// TIA Portal project "Sistema_de_silos" (V16) (continued)
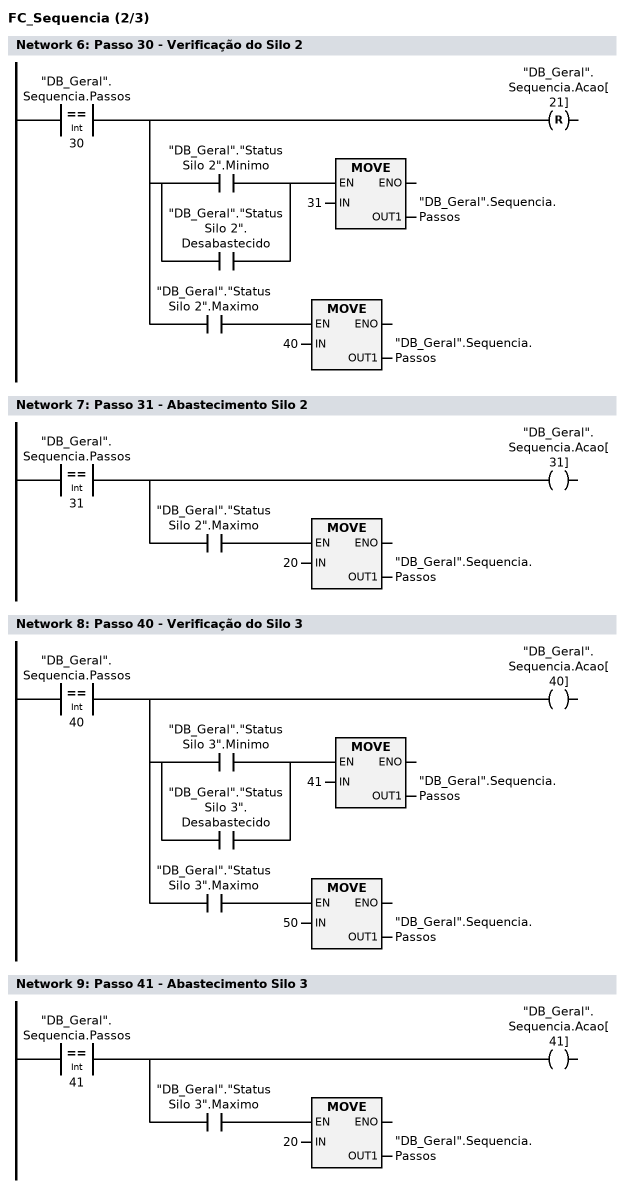
   RUNG wire#powerrail
      { S7_Templates := "SrcType := Int" } EQ_Contact(in1 := "DB_Geral".Sequencia.Passos, in2 := 30)
      wire#w1
      R_Coil( "DB_Geral".Sequencia.Acao[21] )
   END_RUNG
   RUNG wire#w1
      Contact( "DB_Geral"."Status Silo 2".Minimo )
      wire#w2
      Move(in := 31, out1 => "DB_Geral".Sequencia.Passos)
   END_RUNG
   RUNG wire#w1
      Contact( "DB_Geral"."Status Silo 2".Desabastecido )
   END_RUNG wire#w2
   RUNG wire#w1
      Contact( "DB_Geral"."Status Silo 2".Maximo )
      Move(in := 40, out1 => "DB_Geral".Sequencia.Passos)
   END_RUNG
   // the same network as SCL:
   #_w1 := "DB_Geral".Sequencia.Passos = 30;
   IF #_w1 THEN "DB_Geral".Sequencia.Acao[21] := FALSE; END_IF;
   IF #_w1 AND ("DB_Geral"."Status Silo 2".Minimo OR "DB_Geral"."Status Silo 2".Desabastecido) THEN
       "DB_Geral".Sequencia.Passos := 31;
   END_IF;
   IF #_w1 AND "DB_Geral"."Status Silo 2".Maximo THEN "DB_Geral".Sequencia.Passos := 40; END_IF;
END_REGION

REGION Network 7: Passo 31 - Abastecimento Silo 2
   RUNG wire#powerrail
      { S7_Templates := "SrcType := Int" } EQ_Contact(in1 := "DB_Geral".Sequencia.Passos, in2 := 31)
      wire#w1
      Coil( "DB_Geral".Sequencia.Acao[31] )
   END_RUNG
   RUNG wire#w1
      Contact( "DB_Geral"."Status Silo 2".Maximo )
      Move(in := 20, out1 => "DB_Geral".Sequencia.Passos)
   END_RUNG
   // the same network as SCL:
   "DB_Geral".Sequencia.Acao[31] := "DB_Geral".Sequencia.Passos = 31;
   IF ("DB_Geral".Sequencia.Passos = 31) AND "DB_Geral"."Status Silo 2".Maximo THEN
       "DB_Geral".Sequencia.Passos := 20;
   END_IF;
END_REGION

REGION Network 8: Passo 40 - Verificação do Silo 3
   RUNG wire#powerrail
      { S7_Templates := "SrcType := Int" } EQ_Contact(in1 := "DB_Geral".Sequencia.Passos, in2 := 40)
      wire#w1
      Coil( "DB_Geral".Sequencia.Acao[40] )
   END_RUNG
   RUNG wire#w1
      Contact( "DB_Geral"."Status Silo 3".Minimo )
      wire#w2
      Move(in := 41, out1 => "DB_Geral".Sequencia.Passos)
   END_RUNG
   RUNG wire#w1
      Contact( "DB_Geral"."Status Silo 3".Desabastecido )
   END_RUNG wire#w2
   RUNG wire#w1
      Contact( "DB_Geral"."Status Silo 3".Maximo )
      Move(in := 50, out1 => "DB_Geral".Sequencia.Passos)
   END_RUNG
   // the same network as SCL:
   "DB_Geral".Sequencia.Acao[40] := "DB_Geral".Sequencia.Passos = 40;
   #_w1 := "DB_Geral".Sequencia.Passos = 40;
   IF ("DB_Geral".Sequencia.Passos = 40) AND ("DB_Geral"."Status Silo 3".Minimo OR "DB_Geral"."Status Silo 3".Desabastecido) THEN
       "DB_Geral".Sequencia.Passos := 41;
   END_IF;
   IF #_w1 AND "DB_Geral"."Status Silo 3".Maximo THEN "DB_Geral".Sequencia.Passos := 50; END_IF;
END_REGION

REGION Network 9: Passo 41 - Abastecimento Silo 3
   RUNG wire#powerrail
      { S7_Templates := "SrcType := Int" } EQ_Contact(in1 := "DB_Geral".Sequencia.Passos, in2 := 41)
      wire#w1
      Coil( "DB_Geral".Sequencia.Acao[41] )
   END_RUNG
   RUNG wire#w1
      Contact( "DB_Geral"."Status Silo 3".Maximo )
      Move(in := 20, out1 => "DB_Geral".Sequencia.Passos)
   END_RUNG
   // the same network as SCL:
   "DB_Geral".Sequencia.Acao[41] := "DB_Geral".Sequencia.Passos = 41;
   IF ("DB_Geral".Sequencia.Passos = 41) AND "DB_Geral"."Status Silo 3".Maximo THEN
       "DB_Geral".Sequencia.Passos := 20;
   END_IF;
END_REGION

REGION Network 10: Fim de ciclo - Verificação de reserva Maxima do Silo Principal
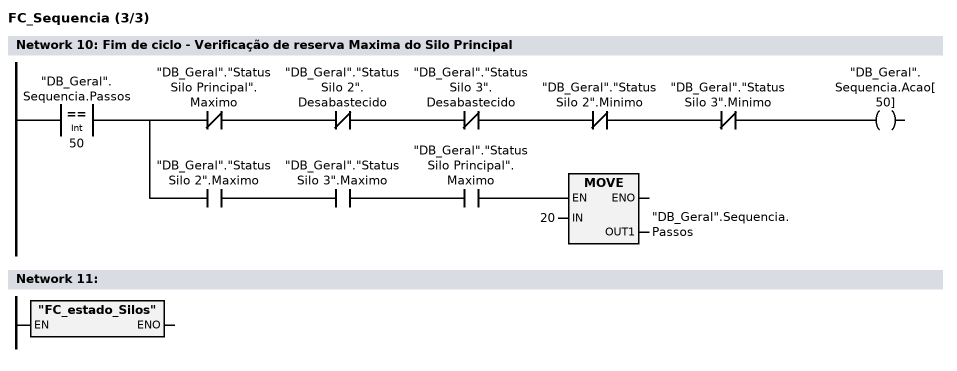
   RUNG wire#powerrail
      { S7_Templates := "SrcType := Int" } EQ_Contact(in1 := "DB_Geral".Sequencia.Passos, in2 := 50)
      wire#w1
      I_Contact( "DB_Geral"."Status Silo Principal".Maximo )
      I_Contact( "DB_Geral"."Status Silo 2".Desabastecido )
      I_Contact( "DB_Geral"."Status Silo 3".Desabastecido )
      I_Contact( "DB_Geral"."Status Silo 2".Minimo )
      I_Contact( "DB_Geral"."Status Silo 3".Minimo )
      Coil( "DB_Geral".Sequencia.Acao[50] )
   END_RUNG
   RUNG wire#w1
      Contact( "DB_Geral"."Status Silo 2".Maximo )
      Contact( "DB_Geral"."Status Silo 3".Maximo )
      Contact( "DB_Geral"."Status Silo Principal".Maximo )
      Move(in := 20, out1 => "DB_Geral".Sequencia.Passos)
   END_RUNG
   // the same network as SCL:
   #_w1 := "DB_Geral".Sequencia.Passos = 50;
   "DB_Geral".Sequencia.Acao[50] := #_w1 AND NOT "DB_Geral"."Status Silo Principal".Maximo AND NOT "DB_Geral"."Status Silo 2".Desabastecido AND NOT "DB_Geral"."Status Silo 3".Desabastecido AND NOT "DB_Geral"."Status Silo 2".Minimo AND NOT "DB_Geral"."Status Silo 3".Minimo;
   IF #_w1 AND "DB_Geral"."Status Silo 2".Maximo AND "DB_Geral"."Status Silo 3".Maximo AND "DB_Geral"."Status Silo Principal".Maximo THEN
       "DB_Geral".Sequencia.Passos := 20;
   END_IF;
END_REGION

REGION Network 11
   RUNG wire#powerrail
      "FC_estado_Silos"()
   END_RUNG
   // the same network as SCL:
   "FC_estado_Silos"();
END_REGION
END_FUNCTION

FUNCTION "FC_Silo_2" : Void   // FC5, LAD
{ S7_Optimized_Access := 'TRUE' }
VERSION : 0.1
   VAR_INPUT
      iAutomatico : Bool;
      iManual : Bool;
      iEmg : Bool;
      iReset : Bool;
      iBtnAbreValvula : Bool;
      iCmdAbreValvula : Bool;
      iCmdAbasteceSilo : Bool;
      iSensorMaximo : Bool;
      iSensorMinimo : Bool;
      iSensorDamper01 : Bool;
      iSensorDamper02 : Bool;
      status_damper : Bool;
      protecao_damper : Bool;
      btnLigaDumper : Bool;
      btnLigaTransportador : Bool;
      iCodinicial : Bool;
   END_VAR
   VAR_IN_OUT
      oAbrirValvula : Bool;
      oLigarDumper : Bool;
      oLigarTransportador : Bool;
      Falha_TimeOut_Desabastecimento : Bool;
      Falha_SensoresNivel : Bool;
      "Status Silo - Minimo" : Bool;
      "Status Silo - Maximo" : Bool;
      "Status Silo - Desabastecido" : Bool;
   END_VAR
   VAR CONSTANT
      Velocidade_fluxo : Int := 12;
   END_VAR
BEGIN

REGION Network 1: Calculo do tempo de vazão - Calculo para fechamento da valvula
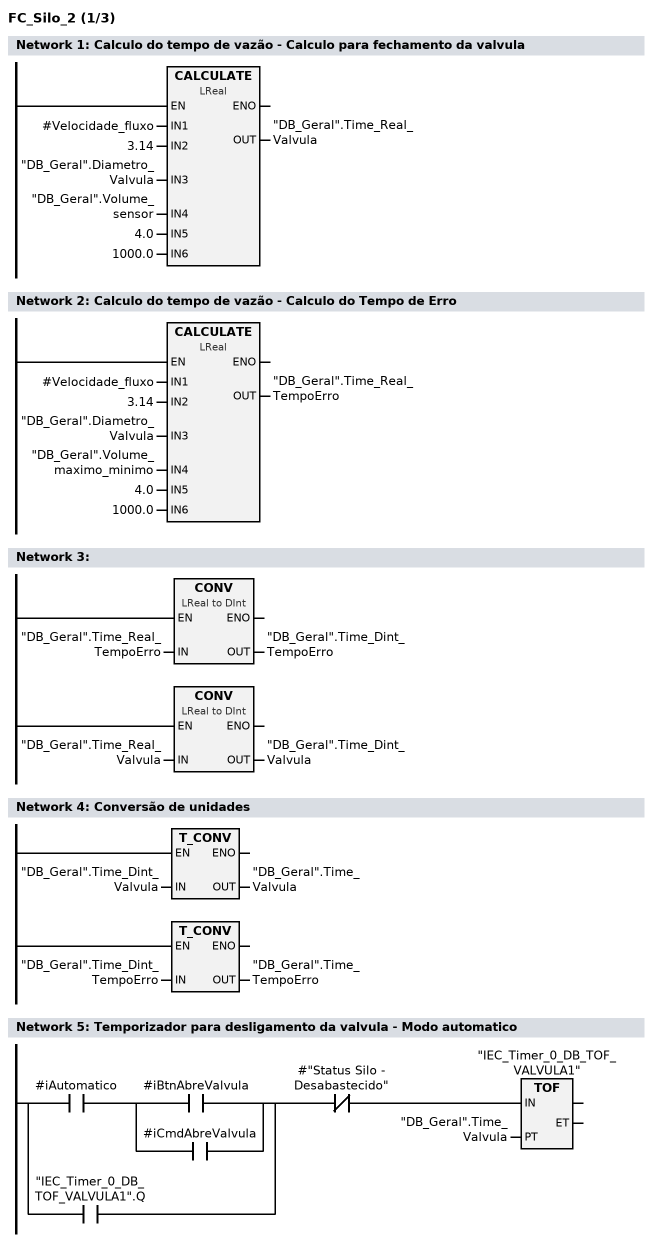
   RUNG wire#powerrail
      { S7_Templates := "SrcType := LReal"; S7_Expression := "(IN4 / (IN1* ((IN2*IN3*IN3) / IN5))) * IN6" } Calculate(in1 := #Velocidade_fluxo, in2 := 3.14, in3 := "DB_Geral".Diametro_Valvula, in4 := "DB_Geral".Volume_sensor, in5 := 4.0, in6 := 1000.0, out => "DB_Geral".Time_Real_Valvula)
   END_RUNG
   // the same network as SCL:
   "DB_Geral".Time_Real_Valvula := ("DB_Geral".Volume_sensor / (#Velocidade_fluxo* ((3.14*"DB_Geral".Diametro_Valvula*"DB_Geral".Diametro_Valvula) / 4.0))) * 1000.0;
END_REGION

REGION Network 2: Calculo do tempo de vazão - Calculo do Tempo de Erro
   RUNG wire#powerrail
      { S7_Templates := "SrcType := LReal"; S7_Expression := "((IN4 / (IN1* ((IN2*IN3*IN3) / IN5))) * IN6)" } Calculate(in1 := #Velocidade_fluxo, in2 := 3.14, in3 := "DB_Geral".Diametro_Valvula, in4 := "DB_Geral".Volume_maximo_minimo, in5 := 4.0, in6 := 1000.0, out => "DB_Geral".Time_Real_TempoErro)
   END_RUNG
   // the same network as SCL:
   "DB_Geral".Time_Real_TempoErro := (("DB_Geral".Volume_maximo_minimo / (#Velocidade_fluxo* ((3.14*"DB_Geral".Diametro_Valvula*"DB_Geral".Diametro_Valvula) / 4.0))) * 1000.0);
END_REGION

REGION Network 3
   RUNG wire#powerrail
      { S7_Templates := "[SrcType := LReal, DestType := DInt]" } Convert(in := "DB_Geral".Time_Real_TempoErro, out => "DB_Geral".Time_Dint_TempoErro)
   END_RUNG
   RUNG wire#powerrail
      { S7_Templates := "[SrcType := LReal, DestType := DInt]" } Convert(in := "DB_Geral".Time_Real_Valvula, out => "DB_Geral".Time_Dint_Valvula)
   END_RUNG
   // the same network as SCL:
   "DB_Geral".Time_Dint_TempoErro := LREAL_TO_DINT("DB_Geral".Time_Real_TempoErro);
   "DB_Geral".Time_Dint_Valvula := LREAL_TO_DINT("DB_Geral".Time_Real_Valvula);
END_REGION

REGION Network 4: Conversão de unidades
   "DB_Geral".Time_Valvula := T_CONV(IN := "DB_Geral".Time_Dint_Valvula);
   "DB_Geral".Time_TempoErro := T_CONV(IN := "DB_Geral".Time_Dint_TempoErro);
END_REGION

REGION Network 5: Temporizador para desligamento da valvula - Modo automatico
   "IEC_Timer_0_DB_TOF_VALVULA1".TOF(IN := ((#iAutomatico AND (#iBtnAbreValvula OR #iCmdAbreValvula)) OR "IEC_Timer_0_DB_TOF_VALVULA1".Q) AND NOT #"Status Silo - Desabastecido",
                           PT := "DB_Geral".Time_Valvula);
END_REGION

REGION Network 6: Acionamento da Valvula
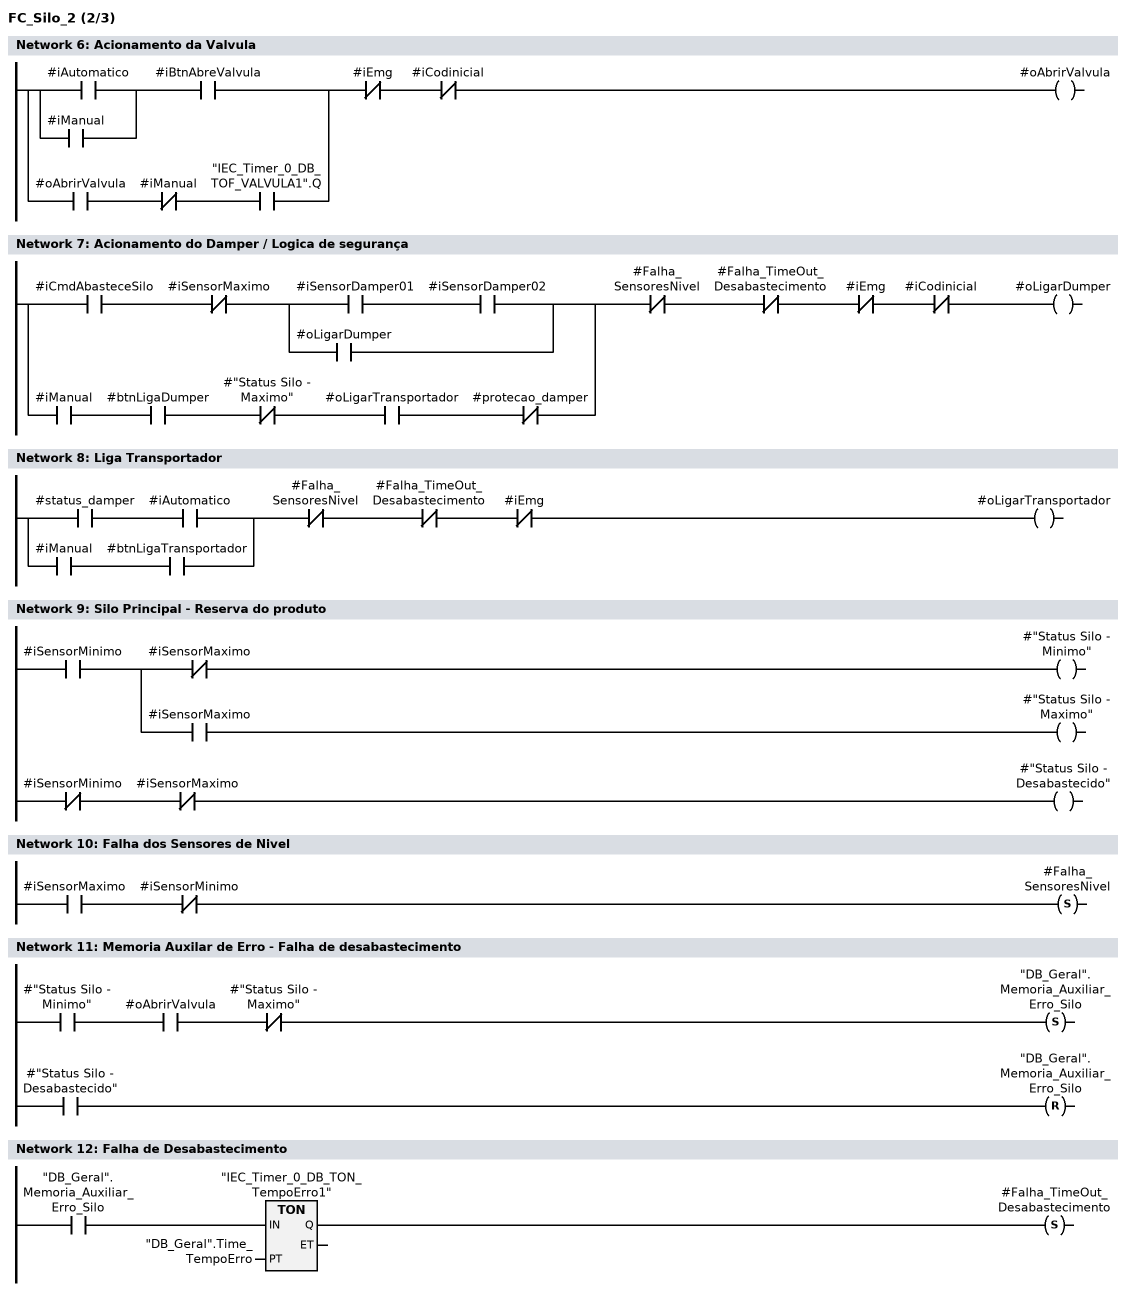
   RUNG wire#powerrail
      Contact( #iAutomatico )
      wire#w1
      Contact( #iBtnAbreValvula )
      wire#w2
      I_Contact( #iEmg )
      I_Contact( #iCodinicial )
      Coil( #oAbrirValvula )
   END_RUNG
   RUNG wire#powerrail
      Contact( #iManual )
   END_RUNG wire#w1
   RUNG wire#powerrail
      Contact( #oAbrirValvula )
      I_Contact( #iManual )
      Contact( "IEC_Timer_0_DB_TOF_VALVULA1".Q )
   END_RUNG wire#w2
   // the same network as SCL:
   #oAbrirValvula := (((#iAutomatico OR #iManual) AND #iBtnAbreValvula) OR (#oAbrirValvula AND NOT #iManual AND "IEC_Timer_0_DB_TOF_VALVULA1".Q)) AND NOT #iEmg AND NOT #iCodinicial;
END_REGION

REGION Network 7: Acionamento do Damper / Logica de segurança
   RUNG wire#powerrail
      Contact( #iCmdAbasteceSilo )
      I_Contact( #iSensorMaximo )
      wire#w1
      Contact( #iSensorDamper01 )
      Contact( #iSensorDamper02 )
      wire#w2
      I_Contact( #Falha_SensoresNivel )
      I_Contact( #Falha_TimeOut_Desabastecimento )
      I_Contact( #iEmg )
      I_Contact( #iCodinicial )
      Coil( #oLigarDumper )
   END_RUNG
   RUNG wire#w1
      Contact( #oLigarDumper )
   END_RUNG wire#w2
   RUNG wire#powerrail
      Contact( #iManual )
      Contact( #btnLigaDumper )
      I_Contact( #"Status Silo - Maximo" )
      Contact( #oLigarTransportador )
      I_Contact( #protecao_damper )
   END_RUNG wire#w2
   // the same network as SCL:
   #oLigarDumper := ((#iCmdAbasteceSilo AND NOT #iSensorMaximo AND ((#iSensorDamper01 AND #iSensorDamper02) OR #oLigarDumper)) OR (#iManual AND #btnLigaDumper AND NOT #"Status Silo - Maximo" AND #oLigarTransportador AND NOT #protecao_damper)) AND NOT #Falha_SensoresNivel AND NOT #Falha_TimeOut_Desabastecimento AND NOT #iEmg AND NOT #iCodinicial;
END_REGION

REGION Network 8: Liga Transportador
   RUNG wire#powerrail
      Contact( #status_damper )
      Contact( #iAutomatico )
      wire#w1
      I_Contact( #Falha_SensoresNivel )
      I_Contact( #Falha_TimeOut_Desabastecimento )
      I_Contact( #iEmg )
      Coil( #oLigarTransportador )
   END_RUNG
   RUNG wire#powerrail
      Contact( #iManual )
      Contact( #btnLigaTransportador )
   END_RUNG wire#w1
   // the same network as SCL:
   #oLigarTransportador := ((#status_damper AND #iAutomatico) OR (#iManual AND #btnLigaTransportador)) AND NOT #Falha_SensoresNivel AND NOT #Falha_TimeOut_Desabastecimento AND NOT #iEmg;
END_REGION

REGION Network 9: Silo Principal - Reserva do produto
   RUNG wire#powerrail
      Contact( #iSensorMinimo )
      wire#w1
      I_Contact( #iSensorMaximo )
      Coil( #"Status Silo - Minimo" )
   END_RUNG
   RUNG wire#w1
      Contact( #iSensorMaximo )
      Coil( #"Status Silo - Maximo" )
   END_RUNG
   RUNG wire#powerrail
      I_Contact( #iSensorMinimo )
      I_Contact( #iSensorMaximo )
      Coil( #"Status Silo - Desabastecido" )
   END_RUNG
   // the same network as SCL:
   #"Status Silo - Minimo" := #iSensorMinimo AND NOT #iSensorMaximo;
   #"Status Silo - Maximo" := #iSensorMinimo AND #iSensorMaximo;
   #"Status Silo - Desabastecido" := NOT #iSensorMinimo AND NOT #iSensorMaximo;
END_REGION

REGION Network 10: Falha dos Sensores de Nivel
   RUNG wire#powerrail
      Contact( #iSensorMaximo )
      I_Contact( #iSensorMinimo )
      S_Coil( #Falha_SensoresNivel )
   END_RUNG
   // the same network as SCL:
   IF #iSensorMaximo AND NOT #iSensorMinimo THEN #Falha_SensoresNivel := TRUE; END_IF;
END_REGION

REGION Network 11: Memoria Auxilar de Erro - Falha de desabastecimento
   RUNG wire#powerrail
      Contact( #"Status Silo - Minimo" )
      Contact( #oAbrirValvula )
      I_Contact( #"Status Silo - Maximo" )
      S_Coil( "DB_Geral".Memoria_Auxiliar_Erro_Silo )
   END_RUNG
   RUNG wire#powerrail
      Contact( #"Status Silo - Desabastecido" )
      R_Coil( "DB_Geral".Memoria_Auxiliar_Erro_Silo )
   END_RUNG
   // the same network as SCL:
   IF #"Status Silo - Minimo" AND #oAbrirValvula AND NOT #"Status Silo - Maximo" THEN
       "DB_Geral".Memoria_Auxiliar_Erro_Silo := TRUE;
   END_IF;
   IF #"Status Silo - Desabastecido" THEN "DB_Geral".Memoria_Auxiliar_Erro_Silo := FALSE; END_IF;
END_REGION

REGION Network 12: Falha de Desabastecimento
   "IEC_Timer_0_DB_TON_TempoErro1".TON(IN := "DB_Geral".Memoria_Auxiliar_Erro_Silo,
                           PT := "DB_Geral".Time_TempoErro);
   IF "IEC_Timer_0_DB_TON_TempoErro1".Q THEN #Falha_TimeOut_Desabastecimento := TRUE; END_IF;
END_REGION

REGION Network 13: Reset - Falhas
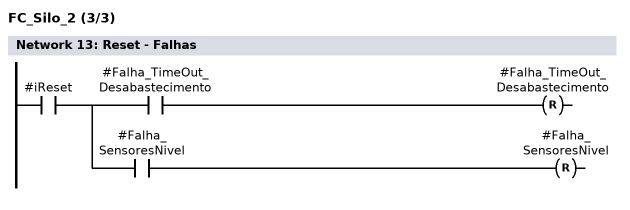
   RUNG wire#powerrail
      Contact( #iReset )
      wire#w1
      Contact( #Falha_TimeOut_Desabastecimento )
      R_Coil( #Falha_TimeOut_Desabastecimento )
   END_RUNG
   RUNG wire#w1
      Contact( #Falha_SensoresNivel )
      R_Coil( #Falha_SensoresNivel )
   END_RUNG
   // the same network as SCL:
   IF #iReset AND #Falha_TimeOut_Desabastecimento THEN #Falha_TimeOut_Desabastecimento := FALSE; END_IF;
   IF #iReset AND #Falha_SensoresNivel THEN #Falha_SensoresNivel := FALSE; END_IF;
END_REGION
END_FUNCTION

FUNCTION "FC_Silo_Principal" : Void   // FC6, LAD
{ S7_Optimized_Access := 'TRUE' }
VERSION : 0.1
   VAR_INPUT
      iAutomatico : Bool;
      iManual : Bool;
      iEmg : Bool;
      iReset : Bool;
      iBtnAbasteceSilo : Bool;
      iCmdAbasteceSilo : Bool;
      iSensorMaximo : Bool;
      iSensorMinimo : Bool;
      iStatusDamper : Bool;
      iCodinicial : Bool;
   END_VAR
   VAR_OUTPUT
      oAbasteceSilo : Bool;
   END_VAR
   VAR_IN_OUT
      Falha_SensoresNivel : Bool;
      "Status Silo - Minimo" : Bool;
      "Status Silo - Maximo" : Bool;
      "Status Silo - Desabastecido" : Bool;
   END_VAR
BEGIN

REGION Network 1
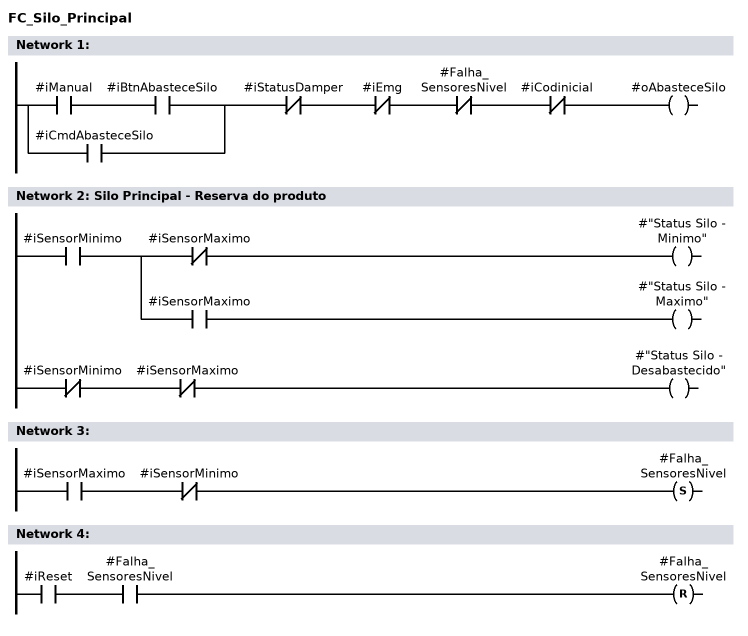
   RUNG wire#powerrail
      Contact( #iManual )
      Contact( #iBtnAbasteceSilo )
      wire#w1
      I_Contact( #iStatusDamper )
      I_Contact( #iEmg )
      I_Contact( #Falha_SensoresNivel )
      I_Contact( #iCodinicial )
      Coil( #oAbasteceSilo )
   END_RUNG
   RUNG wire#powerrail
      Contact( #iCmdAbasteceSilo )
   END_RUNG wire#w1
   // the same network as SCL:
   #oAbasteceSilo := ((#iManual AND #iBtnAbasteceSilo) OR #iCmdAbasteceSilo) AND NOT #iStatusDamper AND NOT #iEmg AND NOT #Falha_SensoresNivel AND NOT #iCodinicial;
END_REGION

REGION Network 2: Silo Principal - Reserva do produto
   RUNG wire#powerrail
      Contact( #iSensorMinimo )
      wire#w1
      I_Contact( #iSensorMaximo )
      Coil( #"Status Silo - Minimo" )
   END_RUNG
   RUNG wire#w1
      Contact( #iSensorMaximo )
      Coil( #"Status Silo - Maximo" )
   END_RUNG
   RUNG wire#powerrail
      I_Contact( #iSensorMinimo )
      I_Contact( #iSensorMaximo )
      Coil( #"Status Silo - Desabastecido" )
   END_RUNG
   // the same network as SCL:
   #"Status Silo - Minimo" := #iSensorMinimo AND NOT #iSensorMaximo;
   #"Status Silo - Maximo" := #iSensorMinimo AND #iSensorMaximo;
   #"Status Silo - Desabastecido" := NOT #iSensorMinimo AND NOT #iSensorMaximo;
END_REGION

REGION Network 3
   RUNG wire#powerrail
      Contact( #iSensorMaximo )
      I_Contact( #iSensorMinimo )
      S_Coil( #Falha_SensoresNivel )
   END_RUNG
   // the same network as SCL:
   IF #iSensorMaximo AND NOT #iSensorMinimo THEN #Falha_SensoresNivel := TRUE; END_IF;
END_REGION

REGION Network 4
   RUNG wire#powerrail
      Contact( #iReset )
      Contact( #Falha_SensoresNivel )
      R_Coil( #Falha_SensoresNivel )
   END_RUNG
   // the same network as SCL:
   IF #iReset AND #Falha_SensoresNivel THEN #Falha_SensoresNivel := FALSE; END_IF;
END_REGION
END_FUNCTION

FUNCTION "FC_Silo_3" : Void   // FC7, LAD
{ S7_Optimized_Access := 'TRUE' }
VERSION : 0.1
   VAR_INPUT
      iAutomatico : Bool;
      iManual : Bool;
      iEmg : Bool;
      iReset : Bool;
      iBtnAbreValvula : Bool;
      iCmdAbreValvula : Bool;
      iCmdAbasteceSilo : Bool;
      iSensorMaximo : Bool;
      iSensorMinimo : Bool;
      iSensorDamper01 : Bool;
      iSensorDamper02 : Bool;
      status_damper : Bool;
      protecao_damper : Bool;
      btnLigaDumper : Bool;
      btnLigaTransportador : Bool;
      iCodinicial : Bool;
   END_VAR
   VAR_IN_OUT
      oAbrirValvula : Bool;
      oLigarDumper : Bool;
      oLigarTransportador : Bool;
      Falha_TimeOut_Desabastecimento : Bool;
      Falha_SensoresNivel : Bool;
      "Status Silo - Minimo" : Bool;
      "Status Silo - Maximo" : Bool;
      "Status Silo - Desabastecido" : Bool;
   END_VAR
   VAR CONSTANT
      Velocidade_fluxo : Int := 12;
   END_VAR
BEGIN

REGION Network 1: Calculo do tempo de vazão - Calculo para fechamento da valvula
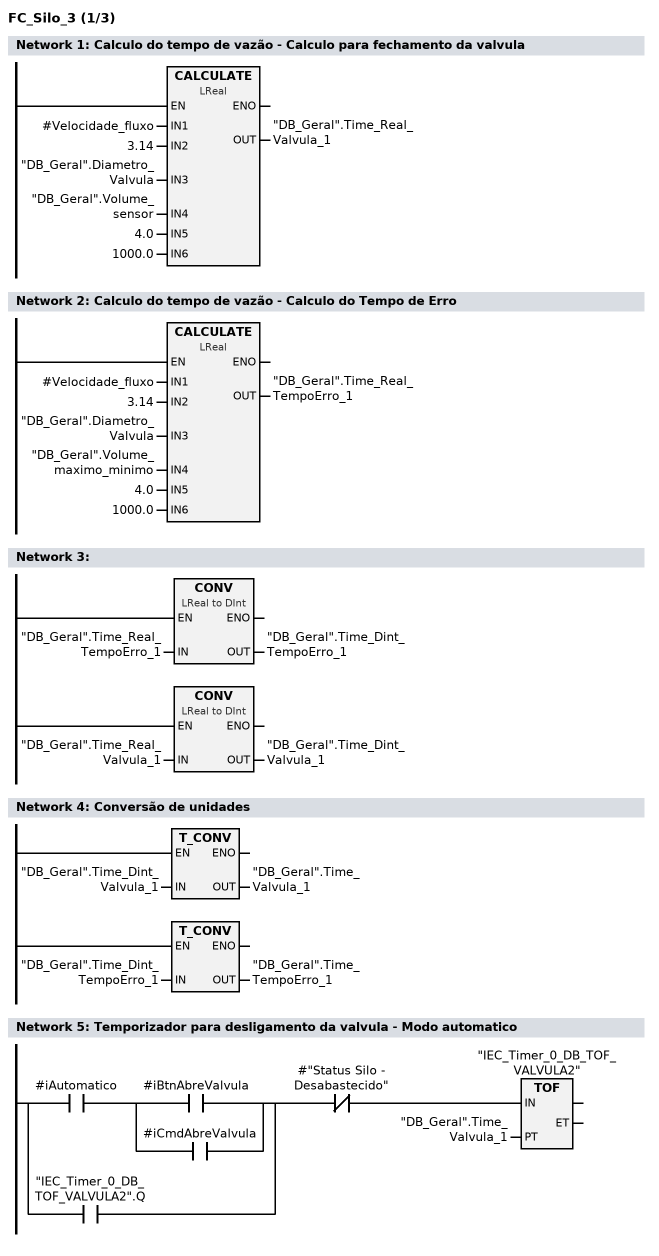
   RUNG wire#powerrail
      { S7_Templates := "SrcType := LReal"; S7_Expression := "(IN4 / (IN1* ((IN2*IN3*IN3) / IN5))) * IN6" } Calculate(in1 := #Velocidade_fluxo, in2 := 3.14, in3 := "DB_Geral".Diametro_Valvula, in4 := "DB_Geral".Volume_sensor, in5 := 4.0, in6 := 1000.0, out => "DB_Geral".Time_Real_Valvula_1)
   END_RUNG
   // the same network as SCL:
   "DB_Geral".Time_Real_Valvula_1 := ("DB_Geral".Volume_sensor / (#Velocidade_fluxo* ((3.14*"DB_Geral".Diametro_Valvula*"DB_Geral".Diametro_Valvula) / 4.0))) * 1000.0;
END_REGION

REGION Network 2: Calculo do tempo de vazão - Calculo do Tempo de Erro
   RUNG wire#powerrail
      { S7_Templates := "SrcType := LReal"; S7_Expression := "(IN4 / (IN1* ((IN2*IN3*IN3) / IN5))) * IN6" } Calculate(in1 := #Velocidade_fluxo, in2 := 3.14, in3 := "DB_Geral".Diametro_Valvula, in4 := "DB_Geral".Volume_maximo_minimo, in5 := 4.0, in6 := 1000.0, out => "DB_Geral".Time_Real_TempoErro_1)
   END_RUNG
   // the same network as SCL:
   "DB_Geral".Time_Real_TempoErro_1 := ("DB_Geral".Volume_maximo_minimo / (#Velocidade_fluxo* ((3.14*"DB_Geral".Diametro_Valvula*"DB_Geral".Diametro_Valvula) / 4.0))) * 1000.0;
END_REGION

REGION Network 3
   RUNG wire#powerrail
      { S7_Templates := "[SrcType := LReal, DestType := DInt]" } Convert(in := "DB_Geral".Time_Real_TempoErro_1, out => "DB_Geral".Time_Dint_TempoErro_1)
   END_RUNG
   RUNG wire#powerrail
      { S7_Templates := "[SrcType := LReal, DestType := DInt]" } Convert(in := "DB_Geral".Time_Real_Valvula_1, out => "DB_Geral".Time_Dint_Valvula_1)
   END_RUNG
   // the same network as SCL:
   "DB_Geral".Time_Dint_TempoErro_1 := LREAL_TO_DINT("DB_Geral".Time_Real_TempoErro_1);
   "DB_Geral".Time_Dint_Valvula_1 := LREAL_TO_DINT("DB_Geral".Time_Real_Valvula_1);
END_REGION

REGION Network 4: Conversão de unidades
   "DB_Geral".Time_Valvula_1 := T_CONV(IN := "DB_Geral".Time_Dint_Valvula_1);
   "DB_Geral".Time_TempoErro_1 := T_CONV(IN := "DB_Geral".Time_Dint_TempoErro_1);
END_REGION

REGION Network 5: Temporizador para desligamento da valvula - Modo automatico
   "IEC_Timer_0_DB_TOF_VALVULA2".TOF(IN := ((#iAutomatico AND (#iBtnAbreValvula OR #iCmdAbreValvula)) OR "IEC_Timer_0_DB_TOF_VALVULA2".Q) AND NOT #"Status Silo - Desabastecido",
                           PT := "DB_Geral".Time_Valvula_1);
END_REGION

REGION Network 6: Acionamento da Valvula
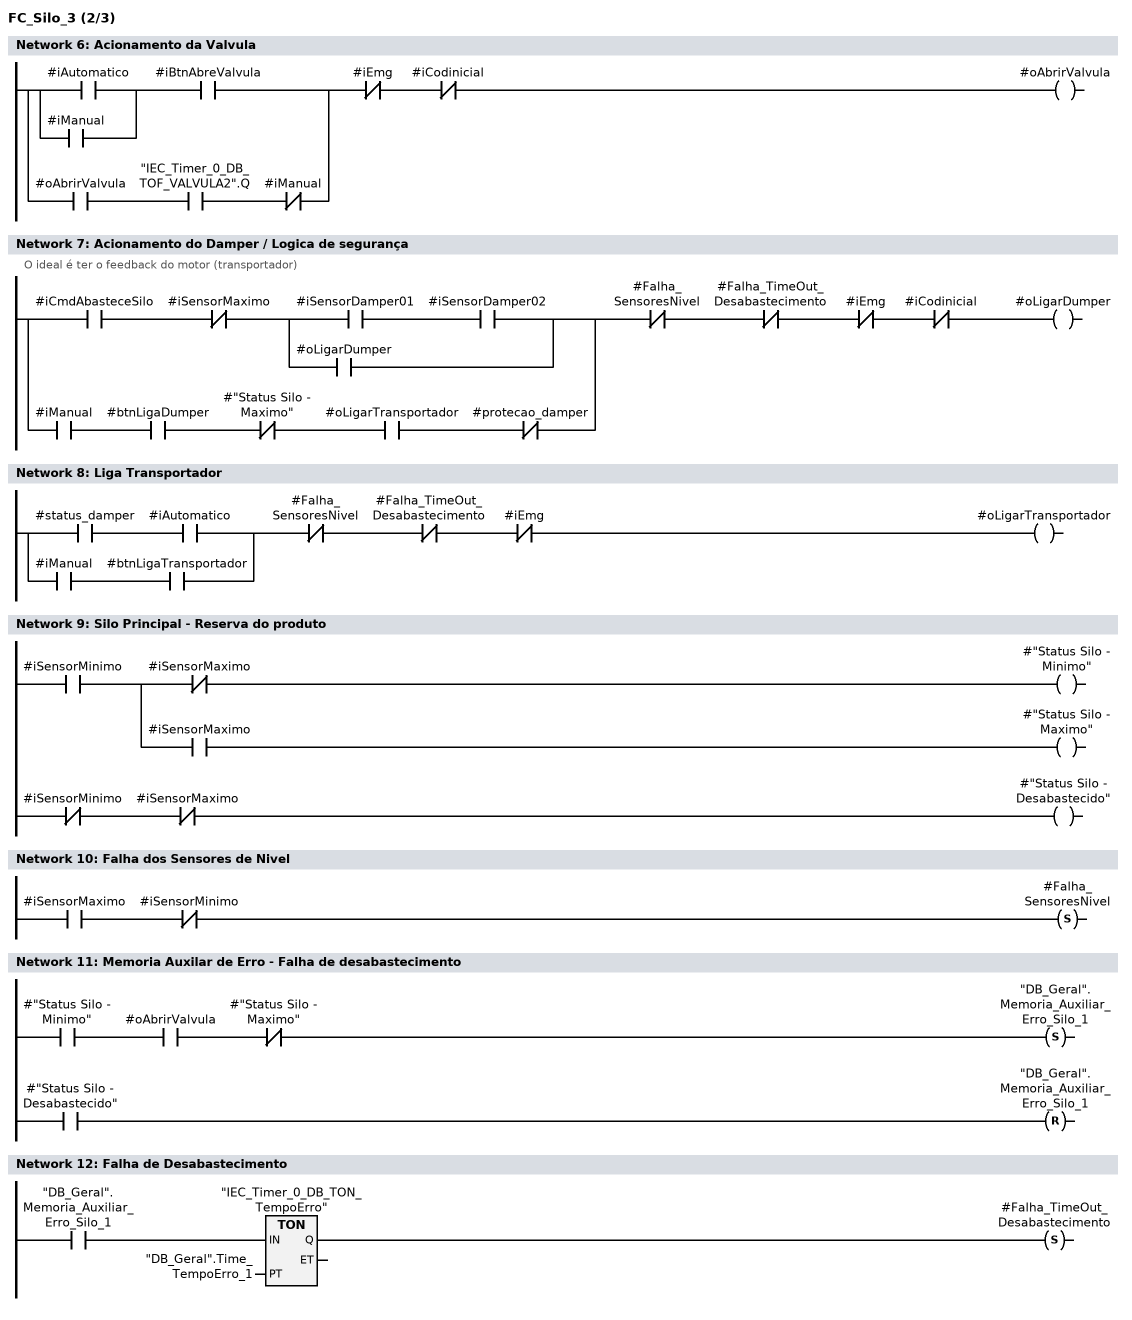
   RUNG wire#powerrail
      Contact( #iAutomatico )
      wire#w1
      Contact( #iBtnAbreValvula )
      wire#w2
      I_Contact( #iEmg )
      I_Contact( #iCodinicial )
      Coil( #oAbrirValvula )
   END_RUNG
   RUNG wire#powerrail
      Contact( #iManual )
   END_RUNG wire#w1
   RUNG wire#powerrail
      Contact( #oAbrirValvula )
      Contact( "IEC_Timer_0_DB_TOF_VALVULA2".Q )
      I_Contact( #iManual )
   END_RUNG wire#w2
   // the same network as SCL:
   #oAbrirValvula := (((#iAutomatico OR #iManual) AND #iBtnAbreValvula) OR (#oAbrirValvula AND "IEC_Timer_0_DB_TOF_VALVULA2".Q AND NOT #iManual)) AND NOT #iEmg AND NOT #iCodinicial;
END_REGION
